
ScreenModuleEditorView "Settings Station Row" 671x200
   TextField "tfLine" at 0,0 size 135x200; Text 'VOLVO 00'
   TextField "tfDropzone" at 135,0 size 40x200; Text '00'
   TextField "tfWIP" at 175,0 size 40x200; Text '00'
   TextField "tfLablBtn00" at 215,0 size 40x25; Text '00'
   TextField "tfAllottedBtn00" at 255,0 size 80x25; Text '00:00'
   TextField "tfCriticalBtn00" at 335,0 size 80x25; Text '00:00'
   TextField "tfPartNumberBtn00" at 415,0 size 256x25; Text '00.00.000.000.0000'
   TextField "tfLablBtn01" at 215,25 size 40x25; Text '00'
   TextField "tfAllottedBtn01" at 255,25 size 80x25; Text '00:00'
   TextField "tfCriticalBtn01" at 335,25 size 80x25; Text '00:00'
   TextField "tfPartNumberBtn01" at 415,25 size 256x25; Text '00.00.000.000.0000'
   TextField "tfLablBtn02" at 215,50 size 40x25; Text '00'
   TextField "tfAllottedBtn02" at 255,50 size 80x25; Text '00:00'
   TextField "tfCriticalBtn02" at 335,50 size 80x25; Text '00:00'
   TextField "tfPartNumberBtn02" at 415,50 size 256x25; Text '00.00.000.000.0000'
   TextField "tfLablBtn03" at 215,75 size 40x25; Text '00'
   TextField "tfAllottedBtn03" at 255,75 size 80x25; Text '00:00'
   TextField "tfCriticalBtn03" at 335,75 size 80x25; Text '00:00'
   TextField "tfPartNumberBtn03" at 415,75 size 256x25; Text '00.00.000.000.0000'
   TextField "tfLablBtn04" at 215,100 size 40x25; Text '00'
   TextField "tfAllottedBtn04" at 255,100 size 80x25; Text '00:00'
   TextField "tfCriticalBtn04" at 335,100 size 80x25; Text '00:00'
   TextField "tfPartNumberBtn04" at 415,100 size 256x25; Text '00.00.000.000.0000'
   TextField "tfLablBtn05" at 215,125 size 40x25; Text '00'
   TextField "tfAllottedBtn05" at 255,125 size 80x25; Text '00:00'
   TextField "tfCriticalBtn05" at 335,125 size 80x25; Text '00:00'
   TextField "tfPartNumberBtn05" at 415,125 size 256x25; Text '00.00.000.000.0000'
   TextField "tfLablBtn06" at 215,150 size 40x25; Text '00'
   TextField "tfAllottedBtn06" at 255,150 size 80x25; Text '00:00'
   TextField "tfCriticalBtn06" at 335,150 size 80x25; Text '00:00'
   TextField "tfPartNumberBtn06" at 415,150 size 256x25; Text '00.00.000.000.0000'
   TextField "tfLablBtn07" at 215,175 size 40x25; Text '00'
   TextField "tfAllottedBtn07" at 255,175 size 80x25; Text '00:00'
   TextField "tfCriticalBtn07" at 335,175 size 80x25; Text '00:00'
   TextField "tfPartNumberBtn07" at 415,175 size 256x25; Text '00.00.000.000.0000'
   TextField "tfPNDoubleBtn00" at 415,0 size 256x25; Text '00.00.000.000.0000 00.00.000.000.0000'
   TextField "tfPNDoubleBtn01" at 415,25 size 256x25; Text '00.00.000.000.0000 00.00.000.000.0000'
   TextField "tfPNDoubleBtn02" at 415,50 size 256x25; Text '00.00.000.000.0000 00.00.000.000.0000'
   TextField "tfPNDoubleBtn03" at 415,75 size 256x25; Text '00.00.000.000.0000 00.00.000.000.0000'
   TextField "tfPNDoubleBtn04" at 415,100 size 256x25; Text '00.00.000.000.0000 00.00.000.000.0000'
   TextField "tfPNDoubleBtn05" at 415,125 size 256x25; Text '00.00.000.000.0000 00.00.000.000.0000'
   TextField "tfPNDoubleBtn06" at 415,150 size 256x25; Text '00.00.000.000.0000 00.00.000.000.0000'
   TextField "tfPNDoubleBtn07" at 415,175 size 256x25; Text '00.00.000.000.0000 00.00.000.000.0000'
*)

(* ===== HMI "HMI_RT_1" =====

graphic list "Top": 0 '100 x 100 Top'; 1 '100 x 100 Actuated Top'

graphic list "Page Up": 0 '100 x 100 Page Up'; 1 '100 x 100 Actuated Page Up'

graphic list "Line Up": 0 '100 x 100 Line Up'; 1 '100 x 100 Actuated Line Up'

graphic list "Line Down": 0 '100 x 100 Line Down'; 1 '100 x 100 Actuated Line Down'

graphic list "Page Down": 0 '100 x 100 Page Down'; 1 '100 x 100 Actuated Page Down'

graphic list "Bottom": 0 '100 x 100 Bottom'; 1 '100 x 100 Actuated Bottom'

ScreenModuleEditorView "Nav Bar: Vertical" 100x600
   Button "btnTop" at 1,1 size 98x98; TextOff 'Text'; PictureList "Top"
   Button "btnPageUp" at 1,101 size 98x98; TextOff 'Text'; PictureList "Page Up"
   Button "btnLineUp" at 1,201 size 98x98; TextOff 'Text'; PictureList "Line Up"
   Button "btnLineDown" at 1,301 size 98x98; TextOff 'Text'; PictureList "Line Down"
   Button "btnPageDown" at 1,401 size 98x98; TextOff 'Text'; PictureList "Page Down"
   Button "btnBottom" at 1,501 size 98x98; TextOff 'Text'; PictureList "Bottom"
*)

(* ===== HMI "HMI_RT_1" =====
system functions are stored by id; their names below are inferred from use

graphic list "Top": 0 '100 x 100 Top'; 1 '100 x 100 Actuated Top'

graphic list "Page Up": 0 '100 x 100 Page Up'; 1 '100 x 100 Actuated Page Up'

graphic list "Line Up": 0 '100 x 100 Line Up'; 1 '100 x 100 Actuated Line Up'

graphic list "Line Down": 0 '100 x 100 Line Down'; 1 '100 x 100 Actuated Line Down'

graphic list "Page Down": 0 '100 x 100 Page Down'; 1 '100 x 100 Actuated Page Down'

graphic list "Bottom": 0 '100 x 100 Bottom'; 1 '100 x 100 Actuated Bottom'

ScreenModuleEditorView "Nav Bar: Vertical" 100x600
   Button "btnTop" at 1,1 size 98x98; TextOff 'Text'; PictureList "Top"
      on Press: SetBit("TableNavBar.top.actuate")
      on Release: ResetBit("TableNavBar.top.actuate")
      Visibility <- "TableNavBar.top.visible"
      ObjectEnable <- "TableNavBar.top.enable"
      ProcessValue <- "TableNavBar.top.listSelect"
      Appearance <- "TableNavBar.top.animate"
   Button "btnPageUp" at 1,101 size 98x98; TextOff 'Text'; PictureList "Page Up"
      on Release: ResetBit("TableNavBar.pageUp.actuate")
      on Press: SetBit("TableNavBar.pageUp.actuate")
      ProcessValue <- "TableNavBar.pageUp.listSelect"
      Appearance <- "TableNavBar.pageUp.animate"
      ObjectEnable <- "TableNavBar.pageUp.enable"
      Visibility <- "TableNavBar.pageUp.visible"
   Button "btnLineUp" at 1,201 size 98x98; TextOff 'Text'; PictureList "Line Up"
      on Release: ResetBit("TableNavBar.lineUp.actuate")
      on Press: SetBit("TableNavBar.lineUp.actuate")
      ProcessValue <- "TableNavBar.lineUp.listSelect"
      Visibility <- "TableNavBar.lineUp.visible"
      ObjectEnable <- "TableNavBar.lineUp.enable"
      Appearance <- "TableNavBar.lineUp.animate"
   Button "btnLineDown" at 1,301 size 98x98; TextOff 'Text'; PictureList "Line Down"
      on Release: ResetBit("TableNavBar.lineDown.actuate")
      on Press: SetBit("TableNavBar.lineDown.actuate")
      ProcessValue <- "TableNavBar.lineDown.listSelect"
      Appearance <- "TableNavBar.lineDown.animate"
      ObjectEnable <- "TableNavBar.lineDown.enable"
      Visibility <- "TableNavBar.lineDown.visible"
   Button "btnPageDown" at 1,401 size 98x98; TextOff 'Text'; PictureList "Page Down"
      on Release: ResetBit("TableNavBar.pageDown.actuate")
      on Press: SetBit("TableNavBar.pageDown.actuate")
      ProcessValue <- "TableNavBar.pageDown.listSelect"
      Visibility <- "TableNavBar.pageDown.visible"
      ObjectEnable <- "TableNavBar.pageDown.enable"
      Appearance <- "TableNavBar.pageDown.animate"
   Button "btnBottom" at 1,501 size 98x98; TextOff 'Text'; PictureList "Bottom"
      on Release: ResetBit("TableNavBar.bottom.actuate")
      on Press: SetBit("TableNavBar.bottom.actuate")
      ProcessValue <- "TableNavBar.bottom.listSelect"
      Appearance <- "TableNavBar.bottom.animate"
      ObjectEnable <- "TableNavBar.bottom.enable"
      Visibility <- "TableNavBar.bottom.visible"
*)

(* ===== HMI "HMI_RT_1" =====
system functions are stored by id; their names below are inferred from use

graphic list "Top": 0 '100 x 100 Top'; 1 '100 x 100 Actuated Top'

graphic list "Page Up": 0 '100 x 100 Page Up'; 1 '100 x 100 Actuated Page Up'

graphic list "Line Up": 0 '100 x 100 Line Up'; 1 '100 x 100 Actuated Line Up'

graphic list "Line Down": 0 '100 x 100 Line Down'; 1 '100 x 100 Actuated Line Down'

graphic list "Page Down": 0 '100 x 100 Page Down'; 1 '100 x 100 Actuated Page Down'

graphic list "Bottom": 0 '100 x 100 Bottom'; 1 '100 x 100 Actuated Bottom'

ScreenModuleEditorView "Nav Bar: Horizontal" 100x600
   Button "btnTop" at 1,1 size 98x98; TextOff 'Text'; PictureList "Top"
      on Release: ResetBit("TableNavBar.top.actuate")
      on Press: SetBit("TableNavBar.top.actuate")
      Visibility <- "TableNavBar.top.visible"
      ObjectEnable <- "TableNavBar.top.enable"
      ProcessValue <- "TableNavBar.top.listSelect"
      Appearance <- "TableNavBar.top.animate"
   Button "btnPageUp" at 1,101 size 98x98; TextOff 'Text'; PictureList "Page Up"
      on Release: ResetBit("TableNavBar.pageUp.actuate")
      on Press: SetBit("TableNavBar.pageUp.actuate")
      Appearance <- "TableNavBar.pageUp.animate"
      ObjectEnable <- "TableNavBar.pageUp.enable"
      ProcessValue <- "TableNavBar.pageUp.listSelect"
      Visibility <- "TableNavBar.pageUp.visible"
   Button "btnLineUp" at 1,201 size 98x98; TextOff 'Text'; PictureList "Line Up"
      on Release: ResetBit("TableNavBar.lineUp.actuate")
      on Press: SetBit("TableNavBar.lineUp.actuate")
      Visibility <- "TableNavBar.lineUp.visible"
      ObjectEnable <- "TableNavBar.lineUp.enable"
      ProcessValue <- "TableNavBar.lineUp.listSelect"
      Appearance <- "TableNavBar.lineUp.animate"
   Button "btnLineDown" at 1,301 size 98x98; TextOff 'Text'; PictureList "Line Down"
      on Release: ResetBit("TableNavBar.lineDown.actuate")
      on Press: SetBit("TableNavBar.lineDown.actuate")
      Appearance <- "TableNavBar.lineDown.animate"
      ObjectEnable <- "TableNavBar.lineDown.enable"
      ProcessValue <- "TableNavBar.lineDown.listSelect"
      Visibility <- "TableNavBar.lineDown.visible"
   Button "btnPageDown" at 1,401 size 98x98; TextOff 'Text'; PictureList "Page Down"
      on Release: ResetBit("TableNavBar.pageDown.actuate")
      on Press: SetBit("TableNavBar.pageDown.actuate")
      Visibility <- "TableNavBar.pageDown.visible"
      ObjectEnable <- "TableNavBar.pageDown.enable"
      ProcessValue <- "TableNavBar.pageDown.listSelect"
      Appearance <- "TableNavBar.pageDown.animate"
   Button "btnBottom" at 1,501 size 98x98; TextOff 'Text'; PictureList "Bottom"
      on Release: ResetBit("TableNavBar.bottom.actuate")
      on Press: SetBit("TableNavBar.bottom.actuate")
      Appearance <- "TableNavBar.bottom.animate"
      ObjectEnable <- "TableNavBar.bottom.enable"
      ProcessValue <- "TableNavBar.bottom.listSelect"
      Visibility <- "TableNavBar.bottom.visible"
*)

(* ===== HMI "HMI_RT_1" =====
system functions are stored by id; their names below are inferred from use

graphic list "Top": 0 '100 x 100 Top'; 1 '100 x 100 Actuated Top'

graphic list "Page Up": 0 '100 x 100 Page Up'; 1 '100 x 100 Actuated Page Up'

graphic list "Line Up": 0 '100 x 100 Line Up'; 1 '100 x 100 Actuated Line Up'

graphic list "Line Down": 0 '100 x 100 Line Down'; 1 '100 x 100 Actuated Line Down'

graphic list "Page Down": 0 '100 x 100 Page Down'; 1 '100 x 100 Actuated Page Down'

graphic list "Bottom": 0 '100 x 100 Bottom'; 1 '100 x 100 Actuated Bottom'

ScreenModuleEditorView "Nav Bar: Horizontal" 600x100
   Button "btnTop" at 1,1 size 98x98; TextOff 'Text'; PictureList "Top"
      on Release: ResetBit("TableNavBar.top.actuate")
      on Press: SetBit("TableNavBar.top.actuate")
      Visibility <- "TableNavBar.top.visible"
      ObjectEnable <- "TableNavBar.top.enable"
      ProcessValue <- "TableNavBar.top.listSelect"
      Appearance <- "TableNavBar.top.animate"
   Button "btnPageUp" at 101,1 size 98x98; TextOff 'Text'; PictureList "Page Up"
      on Release: ResetBit("TableNavBar.pageUp.actuate")
      on Press: SetBit("TableNavBar.pageUp.actuate")
      Appearance <- "TableNavBar.pageUp.animate"
      ObjectEnable <- "TableNavBar.pageUp.enable"
      ProcessValue <- "TableNavBar.pageUp.listSelect"
      Visibility <- "TableNavBar.pageUp.visible"
   Button "btnLineUp" at 201,1 size 98x98; TextOff 'Text'; PictureList "Line Up"
      on Release: ResetBit("TableNavBar.lineUp.actuate")
      on Press: SetBit("TableNavBar.lineUp.actuate")
      Visibility <- "TableNavBar.lineUp.visible"
      ObjectEnable <- "TableNavBar.lineUp.enable"
      ProcessValue <- "TableNavBar.lineUp.listSelect"
      Appearance <- "TableNavBar.lineUp.animate"
   Button "btnLineDown" at 301,1 size 98x98; TextOff 'Text'; PictureList "Line Down"
      on Release: ResetBit("TableNavBar.lineDown.actuate")
      on Press: SetBit("TableNavBar.lineDown.actuate")
      Appearance <- "TableNavBar.lineDown.animate"
      ObjectEnable <- "TableNavBar.lineDown.enable"
      ProcessValue <- "TableNavBar.lineDown.listSelect"
      Visibility <- "TableNavBar.lineDown.visible"
   Button "btnPageDown" at 401,1 size 98x98; TextOff 'Text'; PictureList "Page Down"
      on Release: ResetBit("TableNavBar.pageDown.actuate")
      on Press: SetBit("TableNavBar.pageDown.actuate")
      Visibility <- "TableNavBar.pageDown.visible"
      ObjectEnable <- "TableNavBar.pageDown.enable"
      ProcessValue <- "TableNavBar.pageDown.listSelect"
      Appearance <- "TableNavBar.pageDown.animate"
   Button "btnBottom" at 501,1 size 98x98; TextOff 'Text'; PictureList "Bottom"
      on Release: ResetBit("TableNavBar.bottom.actuate")
      on Press: SetBit("TableNavBar.bottom.actuate")
      Appearance <- "TableNavBar.bottom.animate"
      ObjectEnable <- "TableNavBar.bottom.enable"
      ProcessValue <- "TableNavBar.bottom.listSelect"
      Visibility <- "TableNavBar.bottom.visible"
*)

(* ===== HMI "HMI_RT_1" =====
system functions are stored by id; their names below are inferred from use

ScreenModuleEditorView "PB: Dynamic Text Label" 100x100
   Button "pbActuate" at 0,0 size 100x100; TextOff 'Text'
      on Press: SetBit("Interface.actuate")
      on Release: ResetBit("Interface.actuate")
      ObjectEnable <- "Interface.enable"
      Visibility <- "Interface.visible"
   TextField "tfDisplay" at 0,0 size 100x100; Text 'Text'
      Visibility <- "Interface.visible"
      Appearance <- "Interface.animate"
*)

(* ===== HMI "HMI_RT_1" =====
system functions are stored by id; their names below are inferred from use

ScreenModuleEditorView "PB: Static Text Label" 274x45
   Button "Select All Stations" at 0,0 size 274x45; TextOff 'Text'
      on Press: function_b14e0dd5("Interface.actuate", 0)
      Appearance <- "Interface.animate"
      ObjectEnable <- "Interface.animate"
      Visibility <- "Interface.animate"
*)

(* ===== HMI "HMI_RT_1" =====

ScreenModuleEditorView "Settings Station Row" 671x200
   TextField "tfLine" at 0,0 size 215x200; Text 'Text'
      Appearance <- "Interface.line.animate"
      Visibility <- "Interface.line.visibility"
   TextField "tfLablBtn00" at 215,0 size 40x25; Text '1'
      Appearance <- "Interface.btnRows[0].button.animate"
      Visibility <- "Interface.btnRows[0].button.visibility"
   TextField "tfAllottedBtn00" at 255,0 size 80x25; Text 'Text'
      Appearance <- "Interface.btnRows[0].total.animate"
      Visibility <- "Interface.btnRows[0].total.visibility"
   TextField "tfCriticalBtn00" at 335,0 size 80x25; Text 'Text'
      Appearance <- "Interface.btnRows[0].critical.animate"
      Visibility <- "Interface.btnRows[0].critical.visibility"
   TextField "tfPartNumberBtn00" at 415,0 size 256x25; Text 'Text'
      Appearance <- "Interface.btnRows[0].singlePN.animate"
      Visibility <- "Interface.btnRows[0].singlePN.visibility"
   TextField "tfLablBtn01" at 215,25 size 40x25; Text '2'
      Appearance <- "Interface.btnRows[1].button.animate"
      Visibility <- "Interface.btnRows[1].button.visibility"
   TextField "tfAllottedBtn01" at 255,25 size 80x25; Text 'Text'
      Appearance <- "Interface.btnRows[1].total.animate"
      Visibility <- "Interface.btnRows[1].total.visibility"
   TextField "tfCriticalBtn01" at 335,25 size 80x25; Text 'Text'
      Appearance <- "Interface.btnRows[1].critical.animate"
      Visibility <- "Interface.btnRows[1].critical.visibility"
   TextField "tfPartNumberBtn01" at 415,25 size 256x25; Text 'Text'
      Appearance <- "Interface.btnRows[1].singlePN.animate"
      Visibility <- "Interface.btnRows[1].singlePN.visibility"
   TextField "tfLablBtn02" at 215,50 size 40x25; Text '3'
      Appearance <- "Interface.btnRows[2].button.animate"
      Visibility <- "Interface.btnRows[2].button.visibility"
   TextField "tfAllottedBtn02" at 255,50 size 80x25; Text 'Text'
      Appearance <- "Interface.btnRows[2].total.animate"
      Visibility <- "Interface.btnRows[2].total.visibility"
   TextField "tfCriticalBtn02" at 335,50 size 80x25; Text 'Text'
      Appearance <- "Interface.btnRows[2].critical.animate"
      Visibility <- "Interface.btnRows[2].critical.visibility"
   TextField "tfPartNumberBtn02" at 415,50 size 256x25; Text 'Text'
      Appearance <- "Interface.btnRows[2].singlePN.animate"
      Visibility <- "Interface.btnRows[2].singlePN.visibility"
   TextField "tfLablBtn03" at 215,75 size 40x25; Text '4'
      Appearance <- "Interface.btnRows[3].button.animate"
      Visibility <- "Interface.btnRows[3].button.visibility"
   TextField "tfAllottedBtn03" at 255,75 size 80x25; Text 'Text'
      Appearance <- "Interface.btnRows[3].total.animate"
      Visibility <- "Interface.btnRows[3].total.visibility"
   TextField "tfCriticalBtn03" at 335,75 size 80x25; Text 'Text'
      Appearance <- "Interface.btnRows[3].critical.animate"
      Visibility <- "Interface.btnRows[3].critical.visibility"
   TextField "tfPartNumberBtn03" at 415,75 size 256x25; Text 'Text'
      Appearance <- "Interface.btnRows[3].singlePN.animate"
      Visibility <- "Interface.btnRows[3].singlePN.visibility"
   TextField "tfLablBtn04" at 215,100 size 40x25; Text '5'
      Appearance <- "Interface.btnRows[4].button.animate"
      Visibility <- "Interface.btnRows[4].button.visibility"
   TextField "tfAllottedBtn04" at 255,100 size 80x25; Text 'Text'
      Appearance <- "Interface.btnRows[4].total.animate"
      Visibility <- "Interface.btnRows[4].total.visibility"
   TextField "tfCriticalBtn04" at 335,100 size 80x25; Text 'Text'
      Appearance <- "Interface.btnRows[4].critical.animate"
      Visibility <- "Interface.btnRows[4].critical.visibility"
   TextField "tfPartNumberBtn04" at 415,100 size 256x25; Text 'Text'
      Appearance <- "Interface.btnRows[4].singlePN.animate"
      Visibility <- "Interface.btnRows[4].singlePN.visibility"
   TextField "tfLablBtn05" at 215,125 size 40x25; Text '6'
      Appearance <- "Interface.btnRows[5].button.animate"
      Visibility <- "Interface.btnRows[5].button.visibility"
   TextField "tfAllottedBtn05" at 255,125 size 80x25; Text 'Text'
      Appearance <- "Interface.btnRows[5].total.animate"
      Visibility <- "Interface.btnRows[5].total.visibility"
   TextField "tfCriticalBtn05" at 335,125 size 80x25; Text 'Text'
      Appearance <- "Interface.btnRows[5].critical.animate"
      Visibility <- "Interface.btnRows[5].critical.visibility"
   TextField "tfPartNumberBtn05" at 415,125 size 256x25; Text 'Text'
      Appearance <- "Interface.btnRows[5].singlePN.animate"
      Visibility <- "Interface.btnRows[5].singlePN.visibility"
   TextField "tfLablBtn06" at 215,150 size 40x25; Text '7'
      Appearance <- "Interface.btnRows[6].button.animate"
      Visibility <- "Interface.btnRows[6].button.visibility"
   TextField "tfAllottedBtn06" at 255,150 size 80x25; Text 'Text'
      Appearance <- "Interface.btnRows[6].total.animate"
      Visibility <- "Interface.btnRows[6].total.visibility"
   TextField "tfCriticalBtn06" at 335,150 size 80x25; Text 'Text'
      Appearance <- "Interface.btnRows[6].critical.animate"
      Visibility <- "Interface.btnRows[6].critical.visibility"
   TextField "tfPartNumberBtn06" at 415,150 size 256x25; Text 'Text'
      Appearance <- "Interface.btnRows[6].singlePN.animate"
      Visibility <- "Interface.btnRows[6].singlePN.visibility"
   TextField "tfLablBtn07" at 215,175 size 40x25; Text '8'
      Appearance <- "Interface.btnRows[7].button.animate"
      Visibility <- "Interface.btnRows[7].button.visibility"
   TextField "tfAllottedBtn07" at 255,175 size 80x25; Text 'Text'
      Appearance <- "Interface.btnRows[7].total.animate"
      Visibility <- "Interface.btnRows[7].total.visibility"
   TextField "tfCriticalBtn07" at 335,175 size 80x25; Text 'Text'
      Appearance <- "Interface.btnRows[7].critical.animate"
      Visibility <- "Interface.btnRows[7].critical.visibility"
   TextField "tfPartNumberBtn07" at 415,175 size 256x25; Text 'Text'
      Appearance <- "Interface.btnRows[7].singlePN.animate"
      Visibility <- "Interface.btnRows[7].singlePN.visibility"
   TextField "tfPNDoubleBtn00" at 415,0 size 256x25; Text 'Text'
      Appearance <- "Interface.btnRows[0].doublePN.animate"
      Visibility <- "Interface.btnRows[0].doublePN.visibility"
   TextField "tfPNDoubleBtn01" at 415,25 size 256x25; Text 'Text'
      Appearance <- "Interface.btnRows[1].doublePN.animate"
      Visibility <- "Interface.btnRows[1].doublePN.visibility"
   TextField "tfPNDoubleBtn02" at 415,50 size 256x25; Text 'Text'
      Appearance <- "Interface.btnRows[2].doublePN.animate"
      Visibility <- "Interface.btnRows[2].doublePN.visibility"
   TextField "tfPNDoubleBtn03" at 415,75 size 256x25; Text 'Text'
      Appearance <- "Interface.btnRows[3].doublePN.animate"
      Visibility <- "Interface.btnRows[3].doublePN.visibility"
   TextField "tfPNDoubleBtn04" at 415,100 size 256x25; Text 'Text'
      Appearance <- "Interface.btnRows[4].doublePN.animate"
      Visibility <- "Interface.btnRows[4].doublePN.visibility"
   TextField "tfPNDoubleBtn05" at 415,125 size 256x25; Text 'Text'
      Appearance <- "Interface.btnRows[5].doublePN.animate"
      Visibility <- "Interface.btnRows[5].doublePN.visibility"
   TextField "tfPNDoubleBtn06" at 415,150 size 256x25; Text 'Text'
      Appearance <- "Interface.btnRows[6].doublePN.animate"
      Visibility <- "Interface.btnRows[6].doublePN.visibility"
   TextField "tfPNDoubleBtn07" at 415,175 size 256x25; Text 'Text'
      Appearance <- "Interface.btnRows[7].doublePN.animate"
      Visibility <- "Interface.btnRows[7].doublePN.visibility"
*)

(* ===== HMI "HMI_RT_1" =====
system functions are stored by id; their names below are inferred from use

graphic list "Top": 0 '100 x 100 Top'; 1 '100 x 100 Actuated Top'

graphic list "Page Up": 0 '100 x 100 Page Up'; 1 '100 x 100 Actuated Page Up'

graphic list "Line Up": 0 '100 x 100 Line Up'; 1 '100 x 100 Actuated Line Up'

graphic list "Line Down": 0 '100 x 100 Line Down'; 1 '100 x 100 Actuated Line Down'

graphic list "Page Down": 0 '100 x 100 Page Down'; 1 '100 x 100 Actuated Page Down'

graphic list "Bottom": 0 '100 x 100 Bottom'; 1 '100 x 100 Actuated Bottom'

ScreenModuleEditorView "Nav Bar: Vertical" 100x600
   Button "btnTop" at 1,1 size 98x98; TextOff 'Text'; PictureList "Top"
      on Release: ResetBit("Interface.top.actuate")
      on Press: SetBit("Interface.top.actuate")
      Visibility <- "Interface.top.visible"
      ObjectEnable <- "Interface.top.enable"
      ProcessValue <- "Interface.top.listSelect"
      Appearance <- "Interface.top.animate"
   Button "btnPageUp" at 1,101 size 98x98; TextOff 'Text'; PictureList "Page Up"
      on Release: ResetBit("Interface.pageUp.actuate")
      on Press: SetBit("Interface.pageUp.actuate")
      Appearance <- "Interface.pageUp.animate"
      ObjectEnable <- "Interface.pageUp.enable"
      ProcessValue <- "Interface.pageUp.listSelect"
      Visibility <- "Interface.pageUp.visible"
   Button "btnLineUp" at 1,201 size 98x98; TextOff 'Text'; PictureList "Line Up"
      on Release: ResetBit("Interface.lineUp.actuate")
      on Press: SetBit("Interface.lineUp.actuate")
      Visibility <- "Interface.lineUp.visible"
      ObjectEnable <- "Interface.lineUp.enable"
      ProcessValue <- "Interface.lineUp.listSelect"
      Appearance <- "Interface.lineUp.animate"
   Button "btnLineDown" at 1,301 size 98x98; TextOff 'Text'; PictureList "Line Down"
      on Release: ResetBit("Interface.lineDown.actuate")
      on Press: SetBit("Interface.lineDown.actuate")
      Appearance <- "Interface.lineDown.animate"
      ObjectEnable <- "Interface.lineDown.enable"
      ProcessValue <- "Interface.lineDown.listSelect"
      Visibility <- "Interface.lineDown.visible"
   Button "btnPageDown" at 1,401 size 98x98; TextOff 'Text'; PictureList "Page Down"
      on Release: ResetBit("Interface.pageDown.actuate")
      on Press: SetBit("Interface.pageDown.actuate")
      Visibility <- "Interface.pageDown.visible"
      ObjectEnable <- "Interface.pageDown.enable"
      ProcessValue <- "Interface.pageDown.listSelect"
      Appearance <- "Interface.pageDown.animate"
   Button "btnBottom" at 1,501 size 98x98; TextOff 'Text'; PictureList "Bottom"
      on Release: ResetBit("Interface.bottom.actuate")
      on Press: SetBit("Interface.bottom.actuate")
      Appearance <- "Interface.bottom.animate"
      ObjectEnable <- "Interface.bottom.enable"
      ProcessValue <- "Interface.bottom.listSelect"
      Visibility <- "Interface.bottom.visible"
*)

(* ===== HMI "HMI_RT_1" =====
system functions are stored by id; their names below are inferred from use

graphic list "Top": 0 '100 x 100 Top'; 1 '100 x 100 Actuated Top'

graphic list "Page Up": 0 '100 x 100 Page Up'; 1 '100 x 100 Actuated Page Up'

graphic list "Line Up": 0 '100 x 100 Line Up'; 1 '100 x 100 Actuated Line Up'

graphic list "Line Down": 0 '100 x 100 Line Down'; 1 '100 x 100 Actuated Line Down'

graphic list "Page Down": 0 '100 x 100 Page Down'; 1 '100 x 100 Actuated Page Down'

graphic list "Bottom": 0 '100 x 100 Bottom'; 1 '100 x 100 Actuated Bottom'

ScreenModuleEditorView "Nav Bar: Vertical" 100x600
   Button "btnTop" at 1,1 size 98x98; TextOff 'Text'; PictureList "Top"
      on Release: ResetBit("Interface.top.actuate")
      on Press: SetBit("Interface.top.actuate")
      Visibility <- "Interface.top.visible"
      ObjectEnable <- "Interface.top.enable"
      ProcessValue <- "Interface.top.listSelect"
      Appearance <- "Interface.top.animate"
   Button "btnPageUp" at 1,101 size 98x98; TextOff 'Text'; PictureList "Page Up"
      on Release: ResetBit("Interface.pageUp.actuate")
      on Press: SetBit("Interface.pageUp.actuate")
      Appearance <- "Interface.pageUp.animate"
      ObjectEnable <- "Interface.pageUp.enable"
      ProcessValue <- "Interface.pageUp.listSelect"
      Visibility <- "Interface.pageUp.visible"
   Button "btnLineUp" at 1,201 size 98x98; TextOff 'Text'; PictureList "Line Up"
      on Release: ResetBit("Interface.lineUp.actuate")
      on Press: SetBit("Interface.lineUp.actuate")
      Visibility <- "Interface.lineUp.visible"
      ObjectEnable <- "Interface.lineUp.enable"
      ProcessValue <- "Interface.lineUp.listSelect"
      Appearance <- "Interface.lineUp.animate"
   Button "btnLineDown" at 1,301 size 98x98; TextOff 'Text'; PictureList "Line Down"
      on Release: ResetBit("Interface.lineDown.actuate")
      on Press: SetBit("Interface.lineDown.actuate")
      Appearance <- "Interface.lineDown.animate"
      ObjectEnable <- "Interface.lineDown.enable"
      ProcessValue <- "Interface.lineDown.listSelect"
      Visibility <- "Interface.lineDown.visible"
   Button "btnPageDown" at 1,401 size 98x98; TextOff 'Text'; PictureList "Page Down"
      on Release: ResetBit("Interface.pageDown.actuate")
      on Press: SetBit("Interface.pageDown.actuate")
      Visibility <- "Interface.pageDown.visible"
      ObjectEnable <- "Interface.pageDown.enable"
      ProcessValue <- "Interface.pageDown.listSelect"
      Appearance <- "Interface.pageDown.animate"
   Button "btnBottom" at 1,501 size 98x98; TextOff 'Text'; PictureList "Bottom"
      on Release: ResetBit("Interface.bottom.actuate")
      on Press: SetBit("Interface.bottom.actuate")
      Appearance <- "Interface.bottom.animate"
      ObjectEnable <- "Interface.bottom.enable"
      ProcessValue <- "Interface.bottom.listSelect"
      Visibility <- "Interface.bottom.visible"
*)

(* ===== HMI "HMI_RT_1" =====
system functions are stored by id; their names below are inferred from use

ScreenModuleEditorView "PB: Dynamic Text Label" 100x100
   Button "pbActuate" at 0,0 size 100x100; TextOff 'Text'
      on Release: ResetBit("Interface.actuate")
      on Press: SetBit("Interface.actuate")
      Visibility <- "Interface.visible"
      ObjectEnable <- "Interface.enable"
   TextField "tfDisplay" at 0,0 size 100x100; Text 'Text'
      Visibility <- "Interface.visible"
      Appearance <- "Interface.animate"
*)

(* ===== HMI "HMI_RT_1" =====
system functions are stored by id; their names below are inferred from use

graphic list "Top": 0 '100 x 100 Top'; 1 '100 x 100 Actuated Top'

graphic list "Page Up": 0 '100 x 100 Page Up'; 1 '100 x 100 Actuated Page Up'

graphic list "Line Up": 0 '100 x 100 Line Up'; 1 '100 x 100 Actuated Line Up'

graphic list "Line Down": 0 '100 x 100 Line Down'; 1 '100 x 100 Actuated Line Down'

graphic list "Page Down": 0 '100 x 100 Page Down'; 1 '100 x 100 Actuated Page Down'

graphic list "Bottom": 0 '100 x 100 Bottom'; 1 '100 x 100 Actuated Bottom'

ScreenModuleEditorView "Nav Bar: Horizontal" 600x100
   Button "btnTop" at 1,1 size 98x98; TextOff 'Text'; PictureList "Top"
      on Release: ResetBit("TableNavBar.top.actuate")
      on Press: SetBit("TableNavBar.top.actuate")
      Visibility <- "TableNavBar.top.visible"
      ObjectEnable <- "TableNavBar.top.enable"
      ProcessValue <- "TableNavBar.top.listSelect"
      Appearance <- "TableNavBar.top.animate"
   Button "btnPageUp" at 101,1 size 98x98; TextOff 'Text'; PictureList "Page Up"
      on Release: ResetBit("TableNavBar.pageUp.actuate")
      on Press: SetBit("TableNavBar.pageUp.actuate")
      Appearance <- "TableNavBar.pageUp.animate"
      ObjectEnable <- "TableNavBar.pageUp.enable"
      ProcessValue <- "TableNavBar.pageUp.listSelect"
      Visibility <- "TableNavBar.pageUp.visible"
   Button "btnLineUp" at 201,1 size 98x98; TextOff 'Text'; PictureList "Line Up"
      on Release: ResetBit("TableNavBar.lineUp.actuate")
      on Press: SetBit("TableNavBar.lineUp.actuate")
      Visibility <- "TableNavBar.lineUp.visible"
      ObjectEnable <- "TableNavBar.lineUp.enable"
      ProcessValue <- "TableNavBar.lineUp.listSelect"
      Appearance <- "TableNavBar.lineUp.animate"
   Button "btnLineDown" at 301,1 size 98x98; TextOff 'Text'; PictureList "Line Down"
      on Release: ResetBit("TableNavBar.lineDown.actuate")
      on Press: SetBit("TableNavBar.lineDown.actuate")
      Appearance <- "TableNavBar.lineDown.animate"
      ObjectEnable <- "TableNavBar.lineDown.enable"
      ProcessValue <- "TableNavBar.lineDown.listSelect"
      Visibility <- "TableNavBar.lineDown.visible"
   Button "btnPageDown" at 401,1 size 98x98; TextOff 'Text'; PictureList "Page Down"
      on Release: ResetBit("TableNavBar.pageDown.actuate")
      on Press: SetBit("TableNavBar.pageDown.actuate")
      Visibility <- "TableNavBar.pageDown.visible"
      ObjectEnable <- "TableNavBar.pageDown.enable"
      ProcessValue <- "TableNavBar.pageDown.listSelect"
      Appearance <- "TableNavBar.pageDown.animate"
   Button "btnBottom" at 501,1 size 98x98; TextOff 'Text'; PictureList "Bottom"
      on Release: ResetBit("TableNavBar.bottom.actuate")
      on Press: SetBit("TableNavBar.bottom.actuate")
      Appearance <- "TableNavBar.bottom.animate"
      ObjectEnable <- "TableNavBar.bottom.enable"
      ProcessValue <- "TableNavBar.bottom.listSelect"
      Visibility <- "TableNavBar.bottom.visible"
*)

(* ===== HMI "HMI_RT_1" =====

ScreenModuleEditorView "Settings Station Row" 671x200
   TextField "tfLine" at 0,0 size 215x200; Text 'Text'
      Visibility <- "Interface.line.visibility"
      Appearance <- "Interface.line.animate"
   TextField "tfLablBtn00" at 215,0 size 40x25; Text '1'
      Visibility <- "Interface.btnRows[0].button.visibility"
      Appearance <- "Interface.btnRows[0].button.animate"
   TextField "tfAllottedBtn00" at 255,0 size 80x25; Text 'Text'
      Visibility <- "Interface.btnRows[0].total.visibility"
      Appearance <- "Interface.btnRows[0].total.animate"
   TextField "tfCriticalBtn00" at 335,0 size 80x25; Text 'Text'
      Visibility <- "Interface.btnRows[0].critical.visibility"
      Appearance <- "Interface.btnRows[0].critical.animate"
   TextField "tfPartNumberBtn00" at 415,0 size 256x25; Text 'Text'
      Visibility <- "Interface.btnRows[0].singlePN.visibility"
      Appearance <- "Interface.btnRows[0].singlePN.animate"
   TextField "tfLablBtn01" at 215,25 size 40x25; Text '2'
      Visibility <- "Interface.btnRows[1].button.visibility"
      Appearance <- "Interface.btnRows[1].button.animate"
   TextField "tfAllottedBtn01" at 255,25 size 80x25; Text 'Text'
      Visibility <- "Interface.btnRows[1].total.visibility"
      Appearance <- "Interface.btnRows[1].total.animate"
   TextField "tfCriticalBtn01" at 335,25 size 80x25; Text 'Text'
      Visibility <- "Interface.btnRows[1].critical.visibility"
      Appearance <- "Interface.btnRows[1].critical.animate"
   TextField "tfPartNumberBtn01" at 415,25 size 256x25; Text 'Text'
      Visibility <- "Interface.btnRows[1].singlePN.visibility"
      Appearance <- "Interface.btnRows[1].singlePN.animate"
   TextField "tfLablBtn02" at 215,50 size 40x25; Text '3'
      Visibility <- "Interface.btnRows[2].button.visibility"
      Appearance <- "Interface.btnRows[2].button.animate"
   TextField "tfAllottedBtn02" at 255,50 size 80x25; Text 'Text'
      Visibility <- "Interface.btnRows[2].total.visibility"
      Appearance <- "Interface.btnRows[2].total.animate"
   TextField "tfCriticalBtn02" at 335,50 size 80x25; Text 'Text'
      Visibility <- "Interface.btnRows[2].critical.visibility"
      Appearance <- "Interface.btnRows[2].critical.animate"
   TextField "tfPartNumberBtn02" at 415,50 size 256x25; Text 'Text'
      Visibility <- "Interface.btnRows[2].singlePN.visibility"
      Appearance <- "Interface.btnRows[2].singlePN.animate"
   TextField "tfLablBtn03" at 215,75 size 40x25; Text '4'
      Visibility <- "Interface.btnRows[3].button.visibility"
      Appearance <- "Interface.btnRows[3].button.animate"
   TextField "tfAllottedBtn03" at 255,75 size 80x25; Text 'Text'
      Visibility <- "Interface.btnRows[3].total.visibility"
      Appearance <- "Interface.btnRows[3].total.animate"
   TextField "tfCriticalBtn03" at 335,75 size 80x25; Text 'Text'
      Visibility <- "Interface.btnRows[3].critical.visibility"
      Appearance <- "Interface.btnRows[3].critical.animate"
   TextField "tfPartNumberBtn03" at 415,75 size 256x25; Text 'Text'
      Visibility <- "Interface.btnRows[3].singlePN.visibility"
      Appearance <- "Interface.btnRows[3].singlePN.animate"
   TextField "tfLablBtn04" at 215,100 size 40x25; Text '5'
      Visibility <- "Interface.btnRows[4].button.visibility"
      Appearance <- "Interface.btnRows[4].button.animate"
   TextField "tfAllottedBtn04" at 255,100 size 80x25; Text 'Text'
      Visibility <- "Interface.btnRows[4].total.visibility"
      Appearance <- "Interface.btnRows[4].total.animate"
   TextField "tfCriticalBtn04" at 335,100 size 80x25; Text 'Text'
      Visibility <- "Interface.btnRows[4].critical.visibility"
      Appearance <- "Interface.btnRows[4].critical.animate"
   TextField "tfPartNumberBtn04" at 415,100 size 256x25; Text 'Text'
      Visibility <- "Interface.btnRows[4].singlePN.visibility"
      Appearance <- "Interface.btnRows[4].singlePN.animate"
   TextField "tfLablBtn05" at 215,125 size 40x25; Text '6'
      Visibility <- "Interface.btnRows[5].button.visibility"
      Appearance <- "Interface.btnRows[5].button.animate"
   TextField "tfAllottedBtn05" at 255,125 size 80x25; Text 'Text'
      Visibility <- "Interface.btnRows[5].total.visibility"
      Appearance <- "Interface.btnRows[5].total.animate"
   TextField "tfCriticalBtn05" at 335,125 size 80x25; Text 'Text'
      Visibility <- "Interface.btnRows[5].critical.visibility"
      Appearance <- "Interface.btnRows[5].critical.animate"
   TextField "tfPartNumberBtn05" at 415,125 size 256x25; Text 'Text'
      Visibility <- "Interface.btnRows[5].singlePN.visibility"
      Appearance <- "Interface.btnRows[5].singlePN.animate"
   TextField "tfLablBtn06" at 215,150 size 40x25; Text '7'
      Visibility <- "Interface.btnRows[6].button.visibility"
      Appearance <- "Interface.btnRows[6].button.animate"
   TextField "tfAllottedBtn06" at 255,150 size 80x25; Text 'Text'
      Visibility <- "Interface.btnRows[6].total.visibility"
      Appearance <- "Interface.btnRows[6].total.animate"
   TextField "tfCriticalBtn06" at 335,150 size 80x25; Text 'Text'
      Visibility <- "Interface.btnRows[6].critical.visibility"
      Appearance <- "Interface.btnRows[6].critical.animate"
   TextField "tfPartNumberBtn06" at 415,150 size 256x25; Text 'Text'
      Visibility <- "Interface.btnRows[6].singlePN.visibility"
      Appearance <- "Interface.btnRows[6].singlePN.animate"
   TextField "tfLablBtn07" at 215,175 size 40x25; Text '8'
      Visibility <- "Interface.btnRows[7].button.visibility"
      Appearance <- "Interface.btnRows[7].button.animate"
   TextField "tfAllottedBtn07" at 255,175 size 80x25; Text 'Text'
      Visibility <- "Interface.btnRows[7].total.visibility"
      Appearance <- "Interface.btnRows[7].total.animate"
   TextField "tfCriticalBtn07" at 335,175 size 80x25; Text 'Text'
      Visibility <- "Interface.btnRows[7].critical.visibility"
      Appearance <- "Interface.btnRows[7].critical.animate"
   TextField "tfPartNumberBtn07" at 415,175 size 256x25; Text 'Text'
      Visibility <- "Interface.btnRows[7].singlePN.visibility"
      Appearance <- "Interface.btnRows[7].singlePN.animate"
   TextField "tfPNDoubleBtn00" at 415,0 size 256x25; Text 'Text'
      Visibility <- "Interface.btnRows[0].doublePN.visibility"
      Appearance <- "Interface.btnRows[0].doublePN.animate"
   TextField "tfPNDoubleBtn01" at 415,25 size 256x25; Text 'Text'
      Visibility <- "Interface.btnRows[1].doublePN.visibility"
      Appearance <- "Interface.btnRows[1].doublePN.animate"
   TextField "tfPNDoubleBtn02" at 415,50 size 256x25; Text 'Text'
      Visibility <- "Interface.btnRows[2].doublePN.visibility"
      Appearance <- "Interface.btnRows[2].doublePN.animate"
   TextField "tfPNDoubleBtn03" at 415,75 size 256x25; Text 'Text'
      Visibility <- "Interface.btnRows[3].doublePN.visibility"
      Appearance <- "Interface.btnRows[3].doublePN.animate"
   TextField "tfPNDoubleBtn04" at 415,100 size 256x25; Text 'Text'
      Visibility <- "Interface.btnRows[4].doublePN.visibility"
      Appearance <- "Interface.btnRows[4].doublePN.animate"
   TextField "tfPNDoubleBtn05" at 415,125 size 256x25; Text 'Text'
      Visibility <- "Interface.btnRows[5].doublePN.visibility"
      Appearance <- "Interface.btnRows[5].doublePN.animate"
   TextField "tfPNDoubleBtn06" at 415,150 size 256x25; Text 'Text'
      Visibility <- "Interface.btnRows[6].doublePN.visibility"
      Appearance <- "Interface.btnRows[6].doublePN.animate"
   TextField "tfPNDoubleBtn07" at 415,175 size 256x25; Text 'Text'
      Visibility <- "Interface.btnRows[7].doublePN.visibility"
      Appearance <- "Interface.btnRows[7].doublePN.animate"
*)

(* ===== HMI "HMI_RT_1" =====
system functions are stored by id; their names below are inferred from use

ScreenModuleEditorView "IO Field: Single Width; Stacked" 178x111
   IOField "tfLable" at 0,55 size 178x56; FormatPattern ????????????????????????????????????????
      on OnFinishInput: SetBit("Interface.inputFinished")
      Appearance <- "Interface.animate"
      ProcessValue <- "Interface.value"
      ObjectEnable <- "Interface.enable"
      Visibility <- "Interface.visible"
   TextField "iofData" at 0,0 size 178x55; Text 'Text'
*)

(* ===== HMI "HMI_RT_1" =====
system functions are stored by id; their names below are inferred from use

ScreenModuleEditorView "IO Field: Single Width; Stacked" 178x111
   IOField "tfLable" at 0,55 size 178x56; FormatPattern ????????????????????????????????????????
      on OnFinishInput: SetBit("Interface.inputFinished")
      Appearance <- "Interface.animate"
      Visibility <- "Interface.visible"
      ProcessValue <- "Interface.value"
      ObjectEnable <- "Interface.enable"
   TextField "iofData" at 0,0 size 178x55; Text 'Text'
      Visibility <- "Interface.visible"
*)

(* ===== HMI "HMI_RT_1" =====
system functions are stored by id; their names below are inferred from use

ScreenModuleEditorView "IO Field: Double Width; Stacked" 370x111
   IOField "tfLable" at 0,55 size 370x56; FormatPattern ????????????????????????????????????????
      on OnFinishInput: SetBit("Interface.inputFinished")
      Appearance <- "Interface.animate"
      ProcessValue <- "Interface.value"
      Visibility <- "Interface.visible"
      ObjectEnable <- "Interface.enable"
   TextField "iofData" at 0,0 size 370x55; Text 'Text'
      Visibility <- "Interface.visible"
*)

(* ===== HMI "HMI_RT_1" =====
system functions are stored by id; their names below are inferred from use

ScreenModuleEditorView "PB: Graphic/Text List" 65x45
   Button "Previous Station Group" at 0,0 size 65x45; TextOff 'Text'
      on Press: function_b14e0dd5("Interface.actuate", 0)
      Visibility <- "Interface.animate"
      ObjectEnable <- "Interface.animate"
      Appearance <- "Interface.animate"
*)

(* ===== HMI "HMI_RT_1" =====
system functions are stored by id; their names below are inferred from use

ScreenModuleEditorView "PB: Graphic/Text List" 65x45
   Button "Previous Station Group" at 0,0 size 65x45; TextOff 'Text'
      on Press: function_b14e0dd5("Interface.actuate", 0)
      Visibility <- "Interface.animate"
      ObjectEnable <- "Interface.animate"
      Appearance <- "Interface.animate"
*)

(* ===== HMI "HMI_RT_1" =====
system functions are stored by id; their names below are inferred from use

ScreenModuleEditorView "PB: Station Comm Status (Text Label)" 180x25
   Button "Station Select" at 0,0 size 180x25; TextOff 'Text'
      on Press: function_b14e0dd5("Interface.actuate", 0)
      Appearance <- "Interface.animate"
      ObjectEnable <- "Interface.enable"
      Visibility <- "Interface.visible"
*)

(* ===== HMI "HMI_RT_1" =====
system functions are stored by id; their names below are inferred from use

ScreenModuleEditorView "PB: Graphic/Text List" 65x45
   Button "Previous Station Group" at 0,0 size 65x45; TextOff 'Text'
      on Press: function_b14e0dd5("Interface.actuate", 0)
      Visibility <- "Interface.animate"
      ObjectEnable <- "Interface.animate"
      Appearance <- "Interface.animate"
*)

(* ===== HMI "HMI_RT_1" =====
system functions are stored by id; their names below are inferred from use

graphic list "Top": 0 '100 x 100 Top'; 1 '100 x 100 Actuated Top'

graphic list "Page Up": 0 '100 x 100 Page Up'; 1 '100 x 100 Actuated Page Up'

graphic list "Line Up": 0 '100 x 100 Line Up'; 1 '100 x 100 Actuated Line Up'

graphic list "Line Down": 0 '100 x 100 Line Down'; 1 '100 x 100 Actuated Line Down'

graphic list "Page Down": 0 '100 x 100 Page Down'; 1 '100 x 100 Actuated Page Down'

graphic list "Bottom": 0 '100 x 100 Bottom'; 1 '100 x 100 Actuated Bottom'

ScreenModuleEditorView "Nav Bar: Horizontal" 600x100
   Button "btnTop" at 1,1 size 98x98; TextOff 'Text'; PictureList "Top"
      on Press: function_b14e0dd5("Interface.top.actuate", 0)
      Visibility <- "Interface.top.visible"
      ObjectEnable <- "Interface.top.enable"
      ProcessValue <- "Interface.top.listSelect"
      Appearance <- "Interface.top.animate"
   Button "btnPageUp" at 101,1 size 98x98; TextOff 'Text'; PictureList "Page Up"
      on Press: function_b14e0dd5("Interface.pageUp.actuate", 0)
      Appearance <- "Interface.pageUp.animate"
      ObjectEnable <- "Interface.pageUp.enable"
      ProcessValue <- "Interface.pageUp.listSelect"
      Visibility <- "Interface.pageUp.visible"
   Button "btnLineUp" at 201,1 size 98x98; TextOff 'Text'; PictureList "Line Up"
      on Press: function_b14e0dd5("Interface.lineUp.actuate", 0)
      Visibility <- "Interface.lineUp.visible"
      ObjectEnable <- "Interface.lineUp.enable"
      ProcessValue <- "Interface.lineUp.listSelect"
      Appearance <- "Interface.lineUp.animate"
   Button "btnLineDown" at 301,1 size 98x98; TextOff 'Text'; PictureList "Line Down"
      on Press: function_b14e0dd5("Interface.lineUp.actuate", 0)
      Appearance <- "Interface.lineDown.animate"
      ObjectEnable <- "Interface.lineDown.enable"
      ProcessValue <- "Interface.lineDown.listSelect"
      Visibility <- "Interface.lineDown.visible"
   Button "btnPageDown" at 401,1 size 98x98; TextOff 'Text'; PictureList "Page Down"
      on Press: function_b14e0dd5("Interface.pageDown.actuate", 0)
      Visibility <- "Interface.pageDown.visible"
      ObjectEnable <- "Interface.pageDown.enable"
      ProcessValue <- "Interface.pageDown.listSelect"
      Appearance <- "Interface.pageDown.animate"
   Button "btnBottom" at 501,1 size 98x98; TextOff 'Text'; PictureList "Bottom"
      on Press: function_b14e0dd5("Interface.pageDown.actuate", 0)
      Appearance <- "Interface.bottom.animate"
      ObjectEnable <- "Interface.bottom.enable"
      ProcessValue <- "Interface.bottom.listSelect"
      Visibility <- "Interface.bottom.visible"
*)

(* ===== HMI "HMI_RT_1" =====
system functions are stored by id; their names below are inferred from use

graphic list "Top": 0 '100 x 100 Top'; 1 '100 x 100 Actuated Top'

graphic list "Page Up": 0 '100 x 100 Page Up'; 1 '100 x 100 Actuated Page Up'

graphic list "Line Up": 0 '100 x 100 Line Up'; 1 '100 x 100 Actuated Line Up'

graphic list "Line Down": 0 '100 x 100 Line Down'; 1 '100 x 100 Actuated Line Down'

graphic list "Page Down": 0 '100 x 100 Page Down'; 1 '100 x 100 Actuated Page Down'

graphic list "Bottom": 0 '100 x 100 Bottom'; 1 '100 x 100 Actuated Bottom'

ScreenModuleEditorView "Nav Bar: Horizontal" 600x100
   Button "btnTop" at 1,1 size 98x98; TextOff 'Text'; PictureList "Top"
      on Press: function_b14e0dd5("Interface.top_actuate", 0)
      Appearance <- "Interface.top_animate"
      ObjectEnable <- "Interface.top_enable"
      Visibility <- "Interface.top_visible"
   Button "btnPageUp" at 101,1 size 98x98; TextOff 'Text'; PictureList "Page Up"
      on Press: function_b14e0dd5("Interface.page_up_actuate", 0)
      Visibility <- "Interface.page_up_visible"
      ObjectEnable <- "Interface.page_up_enable"
      Appearance <- "Interface.page_up_animate"
   Button "btnLineUp" at 201,1 size 98x98; TextOff 'Text'; PictureList "Line Up"
      on Press: function_b14e0dd5("Interface.line_up_actuate", 0)
      Visibility <- "Interface.line_up_visible"
      ObjectEnable <- "Interface.line_up_enable"
      Appearance <- "Interface.line_up_animate"
   Button "btnLineDown" at 301,1 size 98x98; TextOff 'Text'; PictureList "Line Down"
      on Press: function_b14e0dd5("Interface.line_down_actuate", 0)
      Appearance <- "Interface.line_down_animate"
      ObjectEnable <- "Interface.line_down_enable"
      Visibility <- "Interface.line_down_visible"
   Button "btnPageDown" at 401,1 size 98x98; TextOff 'Text'; PictureList "Page Down"
      on Press: function_b14e0dd5("Interface.page_down_actuate", 0)
      Visibility <- "Interface.page_down_visible"
      ObjectEnable <- "Interface.page_down_enable"
      Appearance <- "Interface.page_down_animate"
   Button "btnBottom" at 501,1 size 98x98; TextOff 'Text'; PictureList "Bottom"
      on Press: function_b14e0dd5("Interface.botttom_actuate", 0)
      Appearance <- "Interface.botttom_animate"
      ObjectEnable <- "Interface.botttom_enable"
      Visibility <- "Interface.botttom_visible"
*)

(* ===== HMI "HMI_RT_1" =====
system functions are stored by id; their names below are inferred from use

graphic list "Top": 0 '100 x 100 Top'; 1 '100 x 100 Actuated Top'

graphic list "Page Up": 0 '100 x 100 Page Up'; 1 '100 x 100 Actuated Page Up'

graphic list "Line Up": 0 '100 x 100 Line Up'; 1 '100 x 100 Actuated Line Up'

graphic list "Line Down": 0 '100 x 100 Line Down'; 1 '100 x 100 Actuated Line Down'

graphic list "Page Down": 0 '100 x 100 Page Down'; 1 '100 x 100 Actuated Page Down'

graphic list "Bottom": 0 '100 x 100 Bottom'; 1 '100 x 100 Actuated Bottom'

ScreenModuleEditorView "Nav Bar: Vertical" 100x600
   Button "btnTop" at 1,1 size 98x98; TextOff 'Text'; PictureList "Top"
      on Press: function_b14e0dd5("Interface.top_actuate", 0)
      Appearance <- "Interface.top_animate"
      ObjectEnable <- "Interface.top_enable"
      Visibility <- "Interface.top_visible"
   Button "btnPageUp" at 1,101 size 98x98; TextOff 'Text'; PictureList "Page Up"
      on Press: function_b14e0dd5("Interface.page_up_actuate", 0)
      Visibility <- "Interface.page_up_visible"
      ObjectEnable <- "Interface.page_up_enable"
      Appearance <- "Interface.page_up_animate"
   Button "btnLineUp" at 1,201 size 98x98; TextOff 'Text'; PictureList "Line Up"
      on Press: function_b14e0dd5("Interface.line_up_actuate", 0)
      Appearance <- "Interface.line_up_animate"
      ObjectEnable <- "Interface.line_up_enable"
      Visibility <- "Interface.line_up_visible"
   Button "btnLineDown" at 1,301 size 98x98; TextOff 'Text'; PictureList "Line Down"
      on Press: function_b14e0dd5("Interface.line_down_actuate", 0)
      Visibility <- "Interface.line_down_visible"
      ObjectEnable <- "Interface.line_down_enable"
      Appearance <- "Interface.line_down_animate"
   Button "btnPageDown" at 1,401 size 98x98; TextOff 'Text'; PictureList "Page Down"
      on Press: function_b14e0dd5("Interface.page_down_actuate", 0)
      Appearance <- "Interface.page_down_animate"
      ObjectEnable <- "Interface.page_down_enable"
      Visibility <- "Interface.page_down_visible"
   Button "btnBottom" at 1,501 size 98x98; TextOff 'Text'; PictureList "Bottom"
      on Press: SetBit("Interface.bottom_actuate")
      Visibility <- "Interface.bottom_visible"
      ObjectEnable <- "Interface.bottom_enable"
      Appearance <- "Interface.bottom_animate"
*)

(* ===== HMI "HMI_RT_1" =====
system functions are stored by id; their names below are inferred from use

graphic list "Top": 0 '100 x 100 Top'; 1 '100 x 100 Actuated Top'

graphic list "Page Up": 0 '100 x 100 Page Up'; 1 '100 x 100 Actuated Page Up'

graphic list "Line Up": 0 '100 x 100 Line Up'; 1 '100 x 100 Actuated Line Up'

